(* Logix 5000 project; controller NWGG 1756-L72 rev 35.12; software revision 35.00; part 12 of 19 *)
(* tags used below, declared in another part *)
   _101_FEED_AUGER_PIT_101_HM : HOUR_METER;
   _101M : ALIAS FOR O25[9].3;
   _101Y : ALIAS FOR I25[1].3;
   _102_EXPLORE_TANK_41_RECEIVING_LEG_HM : HOUR_METER;
   _102M : ALIAS FOR O25[8].9;
   _102Y : ALIAS FOR I25[0].9;
   _103_TANK_42_RECEIVING_LEG_HM : HOUR_METER;
   _103_TANK_42_RECEIVING_LEG_RUNNING : BOOL;
   _103M : ALIAS FOR O25[8].12;
   _106_TANK_17_AUGER_HM : HOUR_METER;
   _106_TANK_17_AUGER_RUNNING : BOOL;
   _106M : ALIAS FOR O25[9].5;
   _107_SOUTH_BELT_HM : HOUR_METER;
   _107_TANKS_1THRU7_SOUTH_RUNNING : BOOL;
   _107M : ALIAS FOR O25[9].12;
   _108_CENTER_BELT_HM : HOUR_METER;
   _108_CENTER_BELT_RUNNING : BOOL;
   _109_NORTH_BELT_HM : HOUR_METER;
   _109_RAW_RECEIVING_NORTH_BELT_RUNNING : BOOL;
   _110_TANK_16_AUGER_HM : HOUR_METER;
   _110_TANK_16_AUGER_RUNNING : BOOL;
   _111_TANK_17_AUGER_HM : HOUR_METER;
   _111Y : ALIAS FOR I25[1].0;
   _113_HIGHROLLER_TANKS_11TO15_HM : HOUR_METER;
   _113_HIGHROLLER_TANKS_11TO15_RUNNING : BOOL;
   _113_TO_BC1 : ALIAS FOR O25[11].9;
   _113_TO_BC9 : ALIAS FOR O25[11].8;
   _114_TANKS_1THRU7_NORTH_HM : HOUR_METER;
   _114_TANKS_1THRU7_NORTH_RUNNING : BOOL;
   _116_DRAG_16_HM : HOUR_METER;
   _116Y : ALIAS FOR I25[2].10;
   _117_DRAG_17_HM : HOUR_METER;
   _117Y : ALIAS FOR I25[2].8;
   _11_TANK_41_42_HIGHROLLER_HM : HOUR_METER;
   _11_TANK_41_42_HIGHROLLER_RUNNING : BOOL;
   _11M : ALIAS FOR O25[9].2;
   _122_RECIEVING_LEG_HM : HOUR_METER;
   _122M : ALIAS FOR O25[9].1;
   _122Y : ALIAS FOR I25[1].1;
   _123_CLEAN_LEG_HM : HOUR_METER;
   _123_CLEAN_LEG_RUNNING : BOOL;
   _124M : ALIAS FOR O25[9].13;
   _125_COLOR_SORTER_LEG_HM : HOUR_METER;
   _126_ASPERATOR : HOUR_METER;
   _128_SCREENINGS_DRAG_HM : HOUR_METER;
   _1_CLEAN_SEED_UPPER_BELT_HM : HOUR_METER;
   _1_CLEAN_SEED_UPPER_BELT_RUNNING : BOOL;
   _1M : ALIAS FOR O25[9].8;
   _25_16_0 : ALIAS FOR N200[10];
   _25_16_1 : ALIAS FOR N200[11];
   _25_16_2 : ALIAS FOR N200[12];
   _25_16_3 : ALIAS FOR N200[13];
   _2M : ALIAS FOR O25[9].15;
   _35_JUMP_LEG_HM : HOUR_METER;
   _35_JUMP_LEG_RUNNING : BOOL;
   _36_TANK_41_AUGER_HM : HOUR_METER;
   _36_VFD_TO : ALIAS FOR N180[0];
   _36M : ALIAS FOR O25[8].0;
   _36Y : ALIAS FOR I25[0].0;
   _3_LOWER_TANK_CONVAYOR_24TO26_HM : HOUR_METER;
   _3_LOWER_TANK_CONVAYOR_24TO26_RUNNING : BOOL;
   _3_TO_BC5_S : ALIAS FOR O25[11].12;
   _3_TO_BC6_S : ALIAS FOR O25[11].13;
   _42_LOWER_SCREENINGS_DRAG_HM : HOUR_METER;
   _42M : ALIAS FOR O25[11].1;
   _42Y : ALIAS FOR I25[3].1;
   _43_SCREENINGS_LEG_HM : HOUR_METER;
   _43_SCREENINGS_LEG_RUNNING : BOOL;
   _45M : ALIAS FOR O25[8].7;
   _46M : ALIAS FOR O25[8].8;
   _47M : ALIAS FOR O25[9].10;
   _48_CIMBRIA_HM : HOUR_METER;
   _48_VFD_TO : ALIAS FOR N180[2];
   _48M : ALIAS FOR O25[8].3;
   _48Y : ALIAS FOR I25[0].3;
   _49M : ALIAS FOR O25[9].9;
   _4_LOWER_TANK_CONVAYOR_21TO23_HM : HOUR_METER;
   _4_LOWER_TANK_CONVAYOR_21TO23_RUNNING : BOOL;
   _4_TO_BC5_S : ALIAS FOR O25[11].10;
   _4_TO_BC6_S : ALIAS FOR O25[11].11;
   _50M : ALIAS FOR O25[8].14;
   _51_INDENT_HM : HOUR_METER;
   _51_VFD_TO : ALIAS FOR N180[3];
   _51M : ALIAS FOR O25[8].4;
   _51Y : ALIAS FOR I25[0].4;
   _52M : ALIAS FOR O25[8].6;
   _53_VFD_TO : ALIAS FOR N180[1];
   _53M : ALIAS FOR O25[8].2;
   _54M : ALIAS FOR O25[11].3;
   _55M : ALIAS FOR O25[8].1;
   _56M : ALIAS FOR O25[11].2;
   _57M : ALIAS FOR O25[9].6;
   _5_LOWER_CROSS_BELT_HM : HOUR_METER;
   _5Y : ALIAS FOR I25[2].2;
   _701_TRUCK_REVERSING_BELT_HM : HOUR_METER;
   _701_TRUCK_REVERSING_BELT_RUNNING : BOOL;
   _702_CLEAN_JUMP_BELT_HM : HOUR_METER;
   _702Y : ALIAS FOR I25[1].4;
   _703_TREATER_JUMP_BELT_HM : HOUR_METER;
   _703_TREATER_JUMP_BELT_RUNNING : BOOL;
   _9_TREATER_CONVAYOR_HM : HOUR_METER;
   _9_TREATER_CONVAYOR_RUNNING : BOOL;
   ALARM_HORN : ALIAS FOR O25[11].15;
   ALRM_LIGHT : ALIAS FOR O25[11].14;
   Beta : BOOL;
   CLR_SORT_ASP_DELAY : TIMER;
   CLR_SORT_ASPBLR_DELAY : TIMER;
   CLR_SORT_LEG_DELAY : TIMER;
   CLR_SORT_LEG_SPD10 : ALIAS FOR Local:0:I.Data.3;
   CLR_SORT_LEG_SPD20 : ALIAS FOR Local:0:I.Data.4;
   Consumed : DINT;
   hCLR_SORT_LEG_SPD10 : BOOL;
   hCLR_SORT_LEG_SPD20 : BOOL;
   hCLR_SORT_STB : BOOL;
   hCLR_SORT_STRT : BOOL;
   hN_RECVING_PIT_GATE_CLSPB : BOOL;
   hN_RECVING_PIT_GATE_OPNPB : BOOL;
   hSURGE_BIN_HI : BOOL;
   hSURGE_BIN_LO : BOOL;
   I24 : INT[32];
   I25 : INT[32];
   MTR_125_RUNNING : ALIAS FOR Local:0:I.Data.11;
   MTR_125MB : ALIAS FOR Local:5:O.Data.0;
   MTR_126_RUNNING : ALIAS FOR Local:0:I.Data.6;
   MTR_126M : ALIAS FOR Local:5:O.Data.1;
   MTR_126MB : BOOL;
   MTR_127_RUNNING : ALIAS FOR Local:0:I.Data.7;
   MTR_127M : ALIAS FOR Local:5:O.Data.2;
   MTR_127MB : BOOL;
   MTR_128_RUNNING : ALIAS FOR Local:0:I.Data.5;
   MTR_128M : ALIAS FOR Local:5:O.Data.3;
   MTR_128MB : BOOL;
   N180 : DINT[68];
   N190 : DINT[68];
   N27 : DINT[50];
   N_RECVING_PIT_GATE_AUTO : ALIAS FOR Local:0:I.Data.2;
   N_RECVING_PIT_GATE_CLOSE : ALIAS FOR Local:5:O.Data.5;
   N_RECVING_PIT_GATE_OPEN : ALIAS FOR Local:5:O.Data.4;
   O24 : INT[32];
   O25 : INT[32];
   O25_012_Bit00 : ALIAS FOR O25[12].0;
   O25_012_Bit01 : ALIAS FOR O25[12].1;
   O25_012_Bit02 : ALIAS FOR O25[12].2;
   O25_012_Bit03 : ALIAS FOR O25[12].3;
   O25_012_Bit04 : ALIAS FOR O25[12].4;
   O25_012_Bit05 : ALIAS FOR O25[12].5;
   O25_012_Bit06 : ALIAS FOR O25[12].6;
   O25_012_Bit07 : ALIAS FOR O25[12].7;
   O25_012_Bit08 : ALIAS FOR O25[12].8;
   O25_012_Bit09 : ALIAS FOR O25[12].9;
   O25_012_Bit10 : ALIAS FOR O25[12].10;
   O25_012_Bit11 : ALIAS FOR O25[12].11;
   O25_012_Bit12 : ALIAS FOR O25[12].12;
   O25_012_Bit13 : ALIAS FOR O25[12].13;
   O25_012_Bit14 : ALIAS FOR O25[12].14;
   output_Bit : BOOL;
   Output_Bit_2 : BOOL;
   Rack24_1_Mode : BOOL;
   SURGE_BIN_HI : ALIAS FOR Local:0:I.Data.0;
   SURGE_BIN_LO : ALIAS FOR Local:0:I.Data.1;
(* MainProgram, continued *)

ROUTINE Dev_O25_11   (* ladder *)
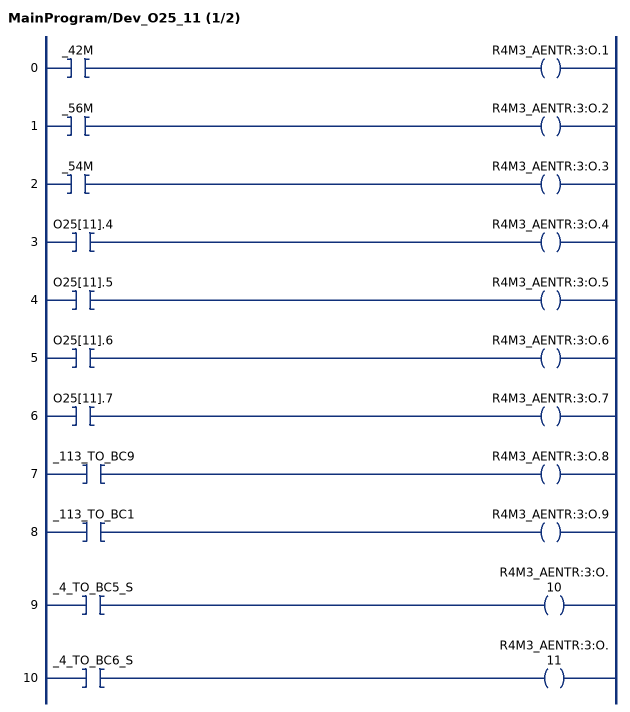
   0: XIC(_42M)OTE(R4M3_AENTR:3:O.1);
   1: XIC(_56M)OTE(R4M3_AENTR:3:O.2);
   2: XIC(_54M)OTE(R4M3_AENTR:3:O.3);
   3: XIC(O25[11].4)OTE(R4M3_AENTR:3:O.4);
   4: XIC(O25[11].5)OTE(R4M3_AENTR:3:O.5);
   5: XIC(O25[11].6)OTE(R4M3_AENTR:3:O.6);
   6: XIC(O25[11].7)OTE(R4M3_AENTR:3:O.7);
   7: XIC(_113_TO_BC9)OTE(R4M3_AENTR:3:O.8);
   8: XIC(_113_TO_BC1)OTE(R4M3_AENTR:3:O.9);
   9: XIC(_4_TO_BC5_S)OTE(R4M3_AENTR:3:O.10);
   10: XIC(_4_TO_BC6_S)OTE(R4M3_AENTR:3:O.11);
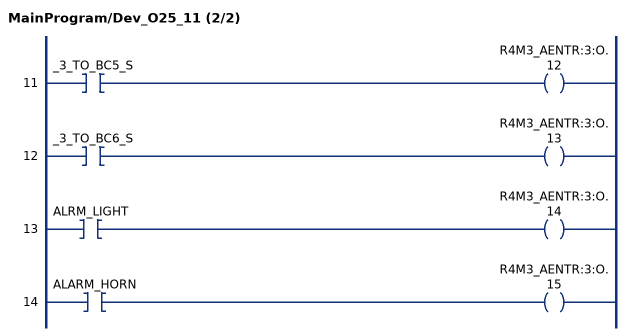
   11: XIC(_3_TO_BC5_S)OTE(R4M3_AENTR:3:O.12);
   12: XIC(_3_TO_BC6_S)OTE(R4M3_AENTR:3:O.13);
   13: XIC(ALRM_LIGHT)OTE(R4M3_AENTR:3:O.14);
   14: XIC(ALARM_HORN)OTE(R4M3_AENTR:3:O.15);
END_ROUTINE

ROUTINE Dev_O25_12   (* ladder *)
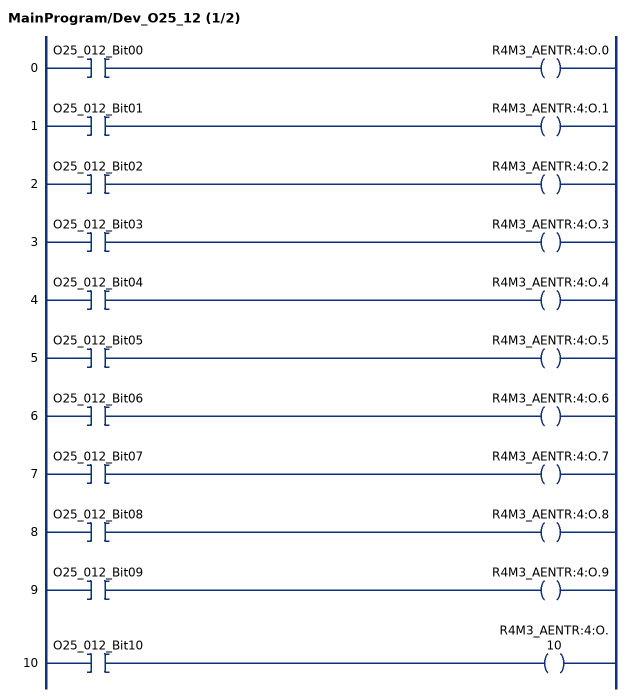
   0: XIC(O25_012_Bit00)OTE(R4M3_AENTR:4:O.0);
   1: XIC(O25_012_Bit01)OTE(R4M3_AENTR:4:O.1);
   2: XIC(O25_012_Bit02)OTE(R4M3_AENTR:4:O.2);
   3: XIC(O25_012_Bit03)OTE(R4M3_AENTR:4:O.3);
   4: XIC(O25_012_Bit04)OTE(R4M3_AENTR:4:O.4);
   5: XIC(O25_012_Bit05)OTE(R4M3_AENTR:4:O.5);
   6: XIC(O25_012_Bit06)OTE(R4M3_AENTR:4:O.6);
   7: XIC(O25_012_Bit07)OTE(R4M3_AENTR:4:O.7);
   8: XIC(O25_012_Bit08)OTE(R4M3_AENTR:4:O.8);
   9: XIC(O25_012_Bit09)OTE(R4M3_AENTR:4:O.9);
   10: XIC(O25_012_Bit10)OTE(R4M3_AENTR:4:O.10);
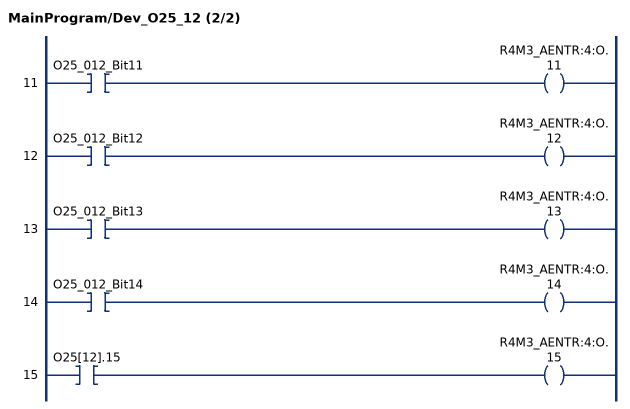
   11: XIC(O25_012_Bit11)OTE(R4M3_AENTR:4:O.11);
   12: XIC(O25_012_Bit12)OTE(R4M3_AENTR:4:O.12);
   13: XIC(O25_012_Bit13)OTE(R4M3_AENTR:4:O.13);
   14: XIC(O25_012_Bit14)OTE(R4M3_AENTR:4:O.14);
   15: XIC(O25[12].15)OTE(R4M3_AENTR:4:O.15);
END_ROUTINE

ROUTINE Dev_O25_8   (* ladder *)
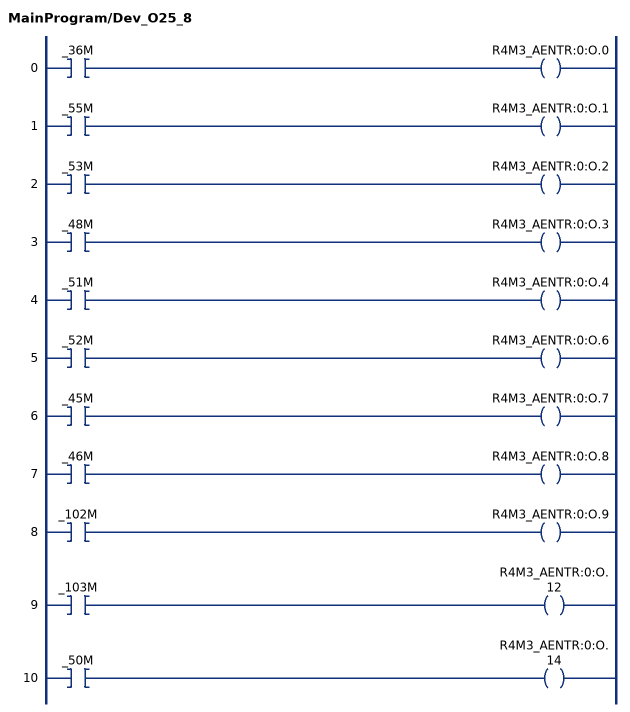
   0: XIC(_36M)OTE(R4M3_AENTR:0:O.0);
   1: XIC(_55M)OTE(R4M3_AENTR:0:O.1);
   2: XIC(_53M)OTE(R4M3_AENTR:0:O.2);
   3: XIC(_48M)OTE(R4M3_AENTR:0:O.3);
   4: XIC(_51M)OTE(R4M3_AENTR:0:O.4);
   5: XIC(_52M)OTE(R4M3_AENTR:0:O.6);
   6: XIC(_45M)OTE(R4M3_AENTR:0:O.7);
   7: XIC(_46M)OTE(R4M3_AENTR:0:O.8);
   8: XIC(_102M)OTE(R4M3_AENTR:0:O.9);
   9: XIC(_103M)OTE(R4M3_AENTR:0:O.12);
   10: XIC(_50M)OTE(R4M3_AENTR:0:O.14);
END_ROUTINE

ROUTINE Dev_O25_9   (* ladder *)
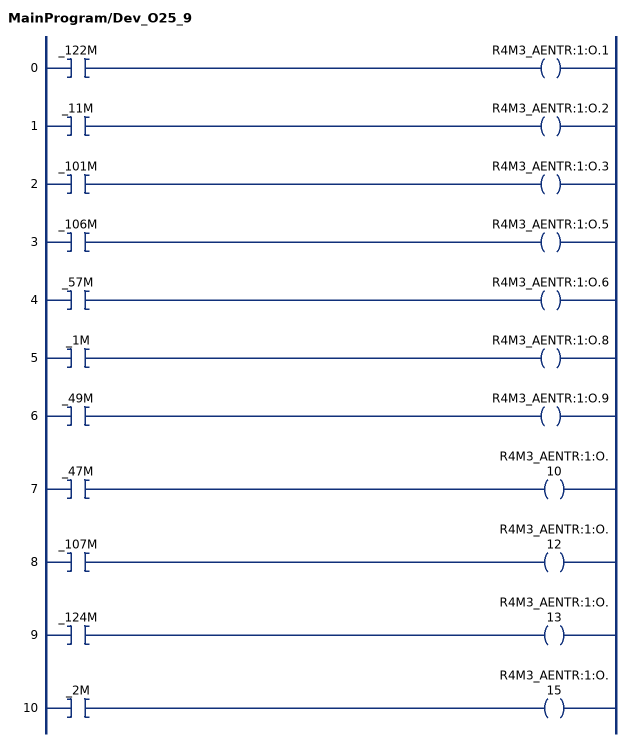
   0: XIC(_122M)OTE(R4M3_AENTR:1:O.1);
   1: XIC(_11M)OTE(R4M3_AENTR:1:O.2);
   2: XIC(_101M)OTE(R4M3_AENTR:1:O.3);
   3: XIC(_106M)OTE(R4M3_AENTR:1:O.5);
   4: XIC(_57M)OTE(R4M3_AENTR:1:O.6);
   5: XIC(_1M)OTE(R4M3_AENTR:1:O.8);
   6: XIC(_49M)OTE(R4M3_AENTR:1:O.9);
   7: XIC(_47M)OTE(R4M3_AENTR:1:O.10);
   8: XIC(_107M)OTE(R4M3_AENTR:1:O.12);
   9: XIC(_124M)OTE(R4M3_AENTR:1:O.13);
   10: XIC(_2M)OTE(R4M3_AENTR:1:O.15);
END_ROUTINE

ROUTINE Disp   (* ladder *)
END_ROUTINE

ROUTINE HOUR_METERS   (* ladder *)
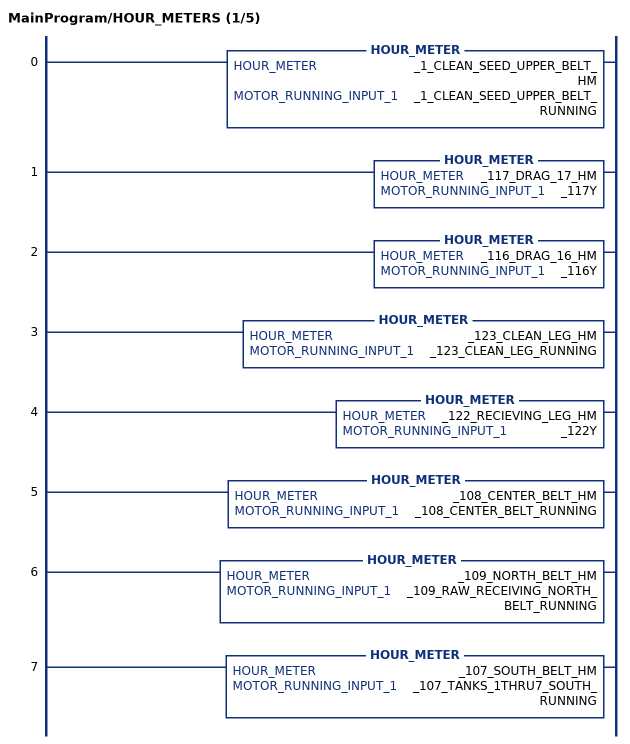
   0: HOUR_METER(_1_CLEAN_SEED_UPPER_BELT_HM,_1_CLEAN_SEED_UPPER_BELT_RUNNING);
   1: HOUR_METER(_117_DRAG_17_HM,_117Y);
   2: HOUR_METER(_116_DRAG_16_HM,_116Y);
   3: HOUR_METER(_123_CLEAN_LEG_HM,_123_CLEAN_LEG_RUNNING);
   4: HOUR_METER(_122_RECIEVING_LEG_HM,_122Y);
   5: HOUR_METER(_108_CENTER_BELT_HM,_108_CENTER_BELT_RUNNING);
   6: HOUR_METER(_109_NORTH_BELT_HM,_109_RAW_RECEIVING_NORTH_BELT_RUNNING);
   7: HOUR_METER(_107_SOUTH_BELT_HM,_107_TANKS_1THRU7_SOUTH_RUNNING);
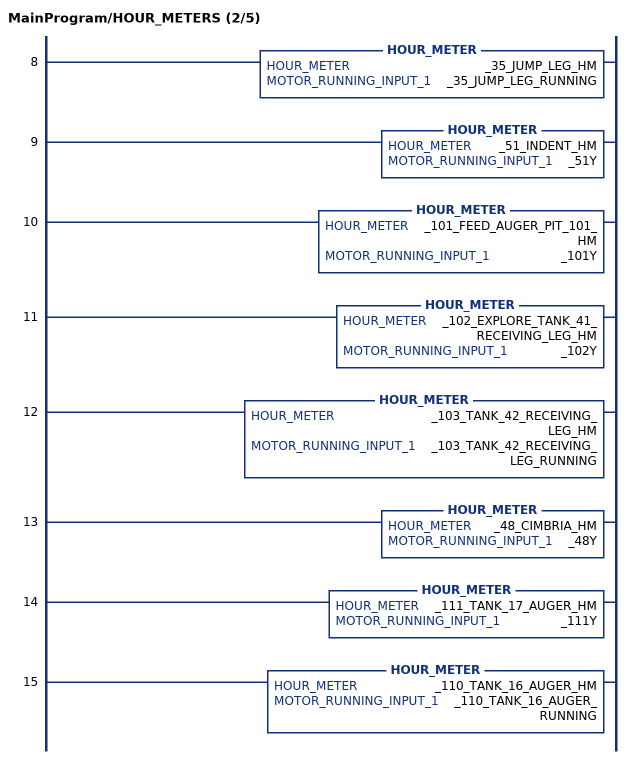
   8: HOUR_METER(_35_JUMP_LEG_HM,_35_JUMP_LEG_RUNNING);
   9: HOUR_METER(_51_INDENT_HM,_51Y);
   10: HOUR_METER(_101_FEED_AUGER_PIT_101_HM,_101Y);
   11: HOUR_METER(_102_EXPLORE_TANK_41_RECEIVING_LEG_HM,_102Y);
   12: HOUR_METER(_103_TANK_42_RECEIVING_LEG_HM,_103_TANK_42_RECEIVING_LEG_RUNNING);
   13: HOUR_METER(_48_CIMBRIA_HM,_48Y);
   14: HOUR_METER(_111_TANK_17_AUGER_HM,_111Y);
   15: HOUR_METER(_110_TANK_16_AUGER_HM,_110_TANK_16_AUGER_RUNNING);
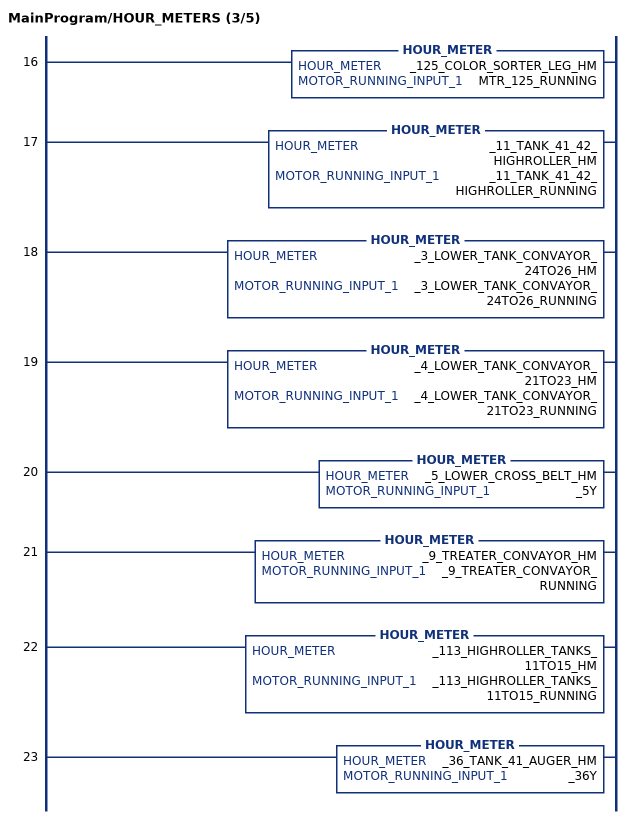
   16: HOUR_METER(_125_COLOR_SORTER_LEG_HM,MTR_125_RUNNING);
   17: HOUR_METER(_11_TANK_41_42_HIGHROLLER_HM,_11_TANK_41_42_HIGHROLLER_RUNNING);
   18: HOUR_METER(_3_LOWER_TANK_CONVAYOR_24TO26_HM,_3_LOWER_TANK_CONVAYOR_24TO26_RUNNING);
   19: HOUR_METER(_4_LOWER_TANK_CONVAYOR_21TO23_HM,_4_LOWER_TANK_CONVAYOR_21TO23_RUNNING);
   20: HOUR_METER(_5_LOWER_CROSS_BELT_HM,_5Y);
   21: HOUR_METER(_9_TREATER_CONVAYOR_HM,_9_TREATER_CONVAYOR_RUNNING);
   22: HOUR_METER(_113_HIGHROLLER_TANKS_11TO15_HM,_113_HIGHROLLER_TANKS_11TO15_RUNNING);
   23: HOUR_METER(_36_TANK_41_AUGER_HM,_36Y);
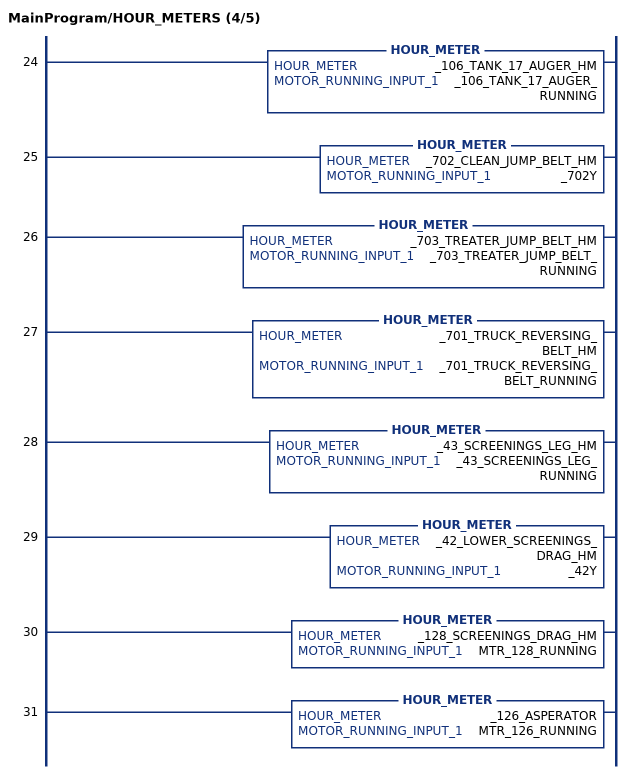
   24: HOUR_METER(_106_TANK_17_AUGER_HM,_106_TANK_17_AUGER_RUNNING);
   25: HOUR_METER(_702_CLEAN_JUMP_BELT_HM,_702Y);
   26: HOUR_METER(_703_TREATER_JUMP_BELT_HM,_703_TREATER_JUMP_BELT_RUNNING);
   27: HOUR_METER(_701_TRUCK_REVERSING_BELT_HM,_701_TRUCK_REVERSING_BELT_RUNNING);
   28: HOUR_METER(_43_SCREENINGS_LEG_HM,_43_SCREENINGS_LEG_RUNNING);
   29: HOUR_METER(_42_LOWER_SCREENINGS_DRAG_HM,_42Y);
   30: HOUR_METER(_128_SCREENINGS_DRAG_HM,MTR_128_RUNNING);
   31: HOUR_METER(_126_ASPERATOR,MTR_126_RUNNING);
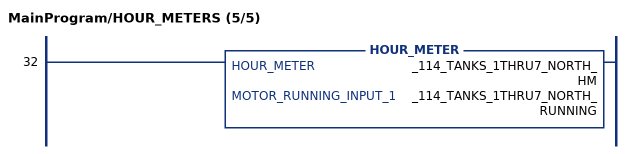
   32: HOUR_METER(_114_TANKS_1THRU7_NORTH_HM,_114_TANKS_1THRU7_NORTH_RUNNING);
END_ROUTINE

ROUTINE MainRoutine   (* ladder *)
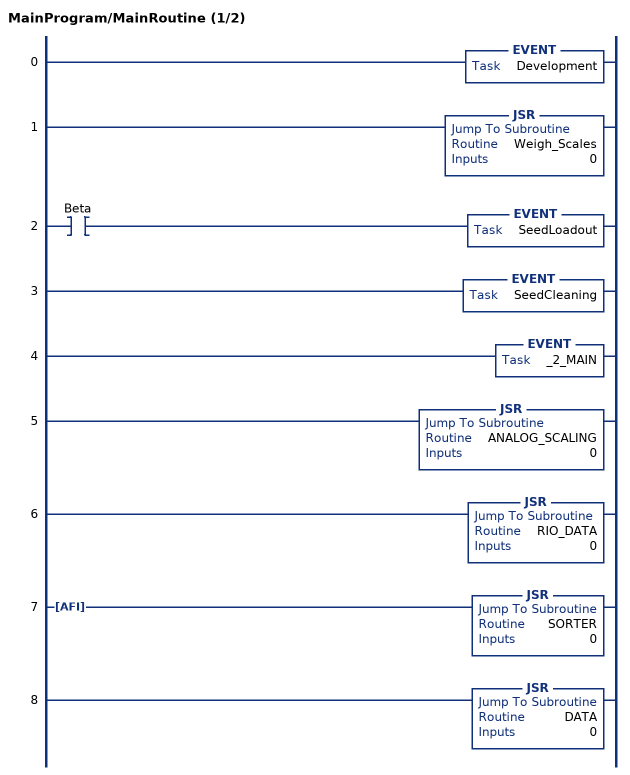
   0: EVENT(Development);
   1: JSR(Weigh_Scales,0);
   2: XIC(Beta)EVENT(SeedLoadout);
   3: EVENT(SeedCleaning);
   4: EVENT(_2_MAIN);
   5: JSR(ANALOG_SCALING,0);
   6: JSR(RIO_DATA,0);
   7: AFI()JSR(SORTER,0);
   8: JSR(DATA,0);
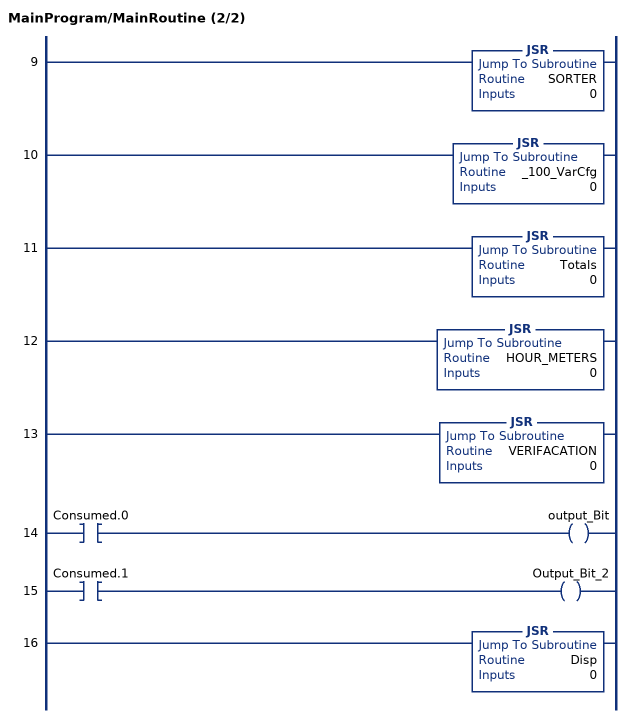
   9: JSR(SORTER,0);
   10: JSR(_100_VarCfg,0);
   11: JSR(Totals,0);
   12: JSR(HOUR_METERS,0);
   13: JSR(VERIFACATION,0);
   14: XIC(Consumed.0)OTE(output_Bit);
   15: XIC(Consumed.1)OTE(Output_Bit_2);
   16: JSR(Disp,0);
END_ROUTINE

ROUTINE RIO_DATA   (* ladder *)
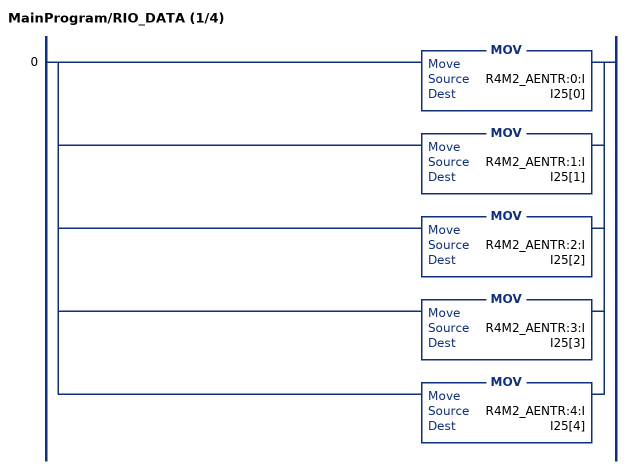
   0: [MOV(R4M2_AENTR:0:I,I25[0]) ,MOV(R4M2_AENTR:1:I,I25[1]) ,MOV(R4M2_AENTR:2:I,I25[2]) ,MOV(R4M2_AENTR:3:I,I25[3]) ,MOV(R4M2_AENTR:4:I,I25[4]) ];
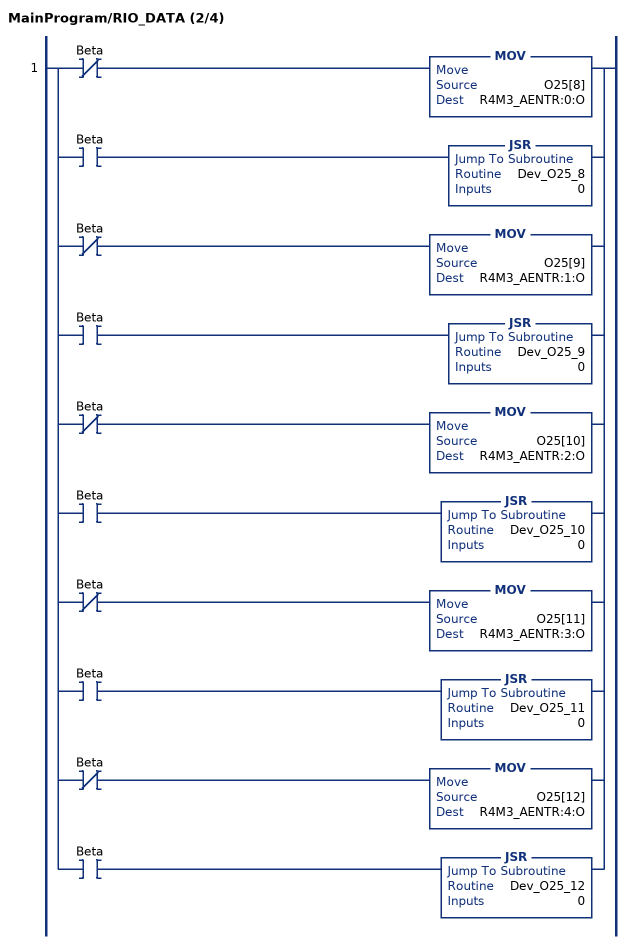
   1: [XIO(Beta) MOV(O25[8],R4M3_AENTR:0:O) ,XIC(Beta) JSR(Dev_O25_8,0) ,XIO(Beta) MOV(O25[9],R4M3_AENTR:1:O) ,XIC(Beta) JSR(Dev_O25_9,0) ,XIO(Beta) MOV(O25[10],R4M3_AENTR:2:O) ,XIC(Beta) JSR(Dev_O25_10,0) ,XIO(Beta) MOV(O25[11],R4M3_AENTR:3:O) ,XIC(Beta) JSR(Dev_O25_11,0) ,XIO(Beta) MOV(O25[12],R4M3_AENTR:4:O) ,XIC(Beta) JSR(Dev_O25_12,0) ];
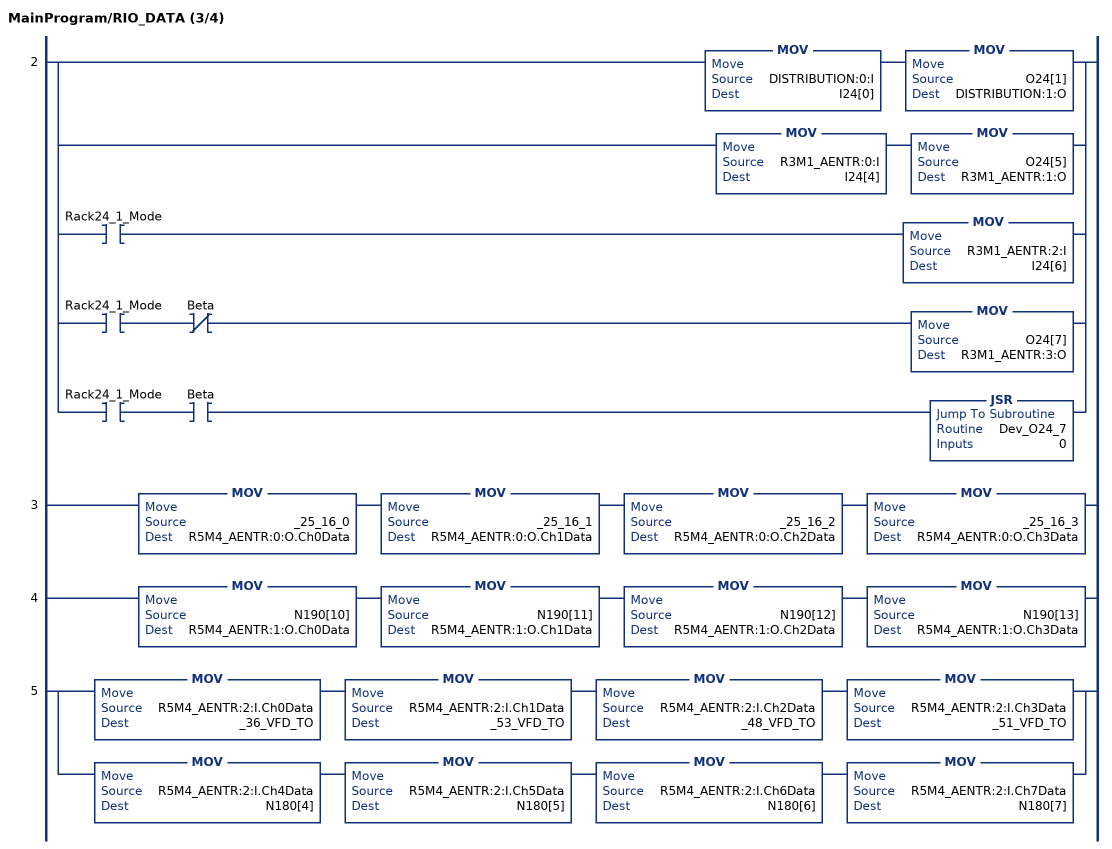
   2: [MOV(DISTRIBUTION:0:I,I24[0]) MOV(O24[1],DISTRIBUTION:1:O) ,MOV(R3M1_AENTR:0:I,I24[4]) MOV(O24[5],R3M1_AENTR:1:O) ,XIC(Rack24_1_Mode) MOV(R3M1_AENTR:2:I,I24[6]) ,XIC(Rack24_1_Mode) XIO(Beta) MOV(O24[7],R3M1_AENTR:3:O) ,XIC(Rack24_1_Mode) XIC(Beta) JSR(Dev_O24_7,0) ];
   3: MOV(_25_16_0,R5M4_AENTR:0:O.Ch0Data)MOV(_25_16_1,R5M4_AENTR:0:O.Ch1Data)MOV(_25_16_2,R5M4_AENTR:0:O.Ch2Data)MOV(_25_16_3,R5M4_AENTR:0:O.Ch3Data);
   4: MOV(N190[10],R5M4_AENTR:1:O.Ch0Data)MOV(N190[11],R5M4_AENTR:1:O.Ch1Data)MOV(N190[12],R5M4_AENTR:1:O.Ch2Data)MOV(N190[13],R5M4_AENTR:1:O.Ch3Data);
   5: [MOV(R5M4_AENTR:2:I.Ch0Data,_36_VFD_TO) MOV(R5M4_AENTR:2:I.Ch1Data,_53_VFD_TO) MOV(R5M4_AENTR:2:I.Ch2Data,_48_VFD_TO) MOV(R5M4_AENTR:2:I.Ch3Data,_51_VFD_TO) ,MOV(R5M4_AENTR:2:I.Ch4Data,N180[4]) MOV(R5M4_AENTR:2:I.Ch5Data,N180[5]) MOV(R5M4_AENTR:2:I.Ch6Data,N180[6]) MOV(R5M4_AENTR:2:I.Ch7Data,N180[7]) ];
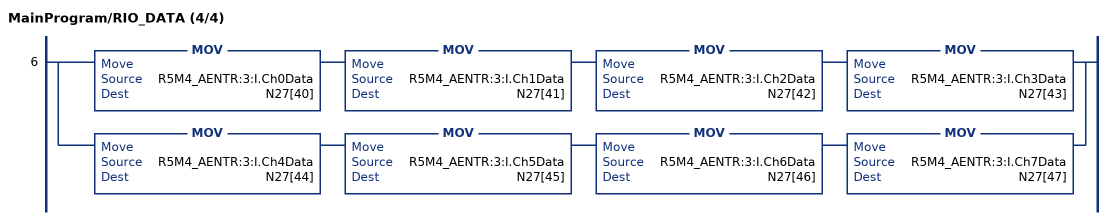
   6: [MOV(R5M4_AENTR:3:I.Ch0Data,N27[40]) MOV(R5M4_AENTR:3:I.Ch1Data,N27[41]) MOV(R5M4_AENTR:3:I.Ch2Data,N27[42]) MOV(R5M4_AENTR:3:I.Ch3Data,N27[43]) ,MOV(R5M4_AENTR:3:I.Ch4Data,N27[44]) MOV(R5M4_AENTR:3:I.Ch5Data,N27[45]) MOV(R5M4_AENTR:3:I.Ch6Data,N27[46]) MOV(R5M4_AENTR:3:I.Ch7Data,N27[47]) ];
END_ROUTINE

ROUTINE SORTER   (* ladder *)
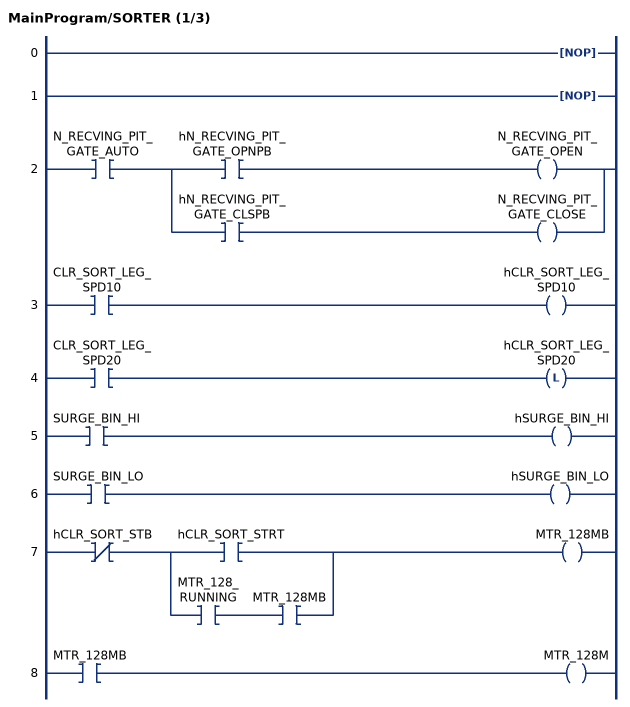
   0: NOP();
   1: NOP();
   2: XIC(N_RECVING_PIT_GATE_AUTO)[XIC(hN_RECVING_PIT_GATE_OPNPB) OTE(N_RECVING_PIT_GATE_OPEN) ,XIC(hN_RECVING_PIT_GATE_CLSPB) OTE(N_RECVING_PIT_GATE_CLOSE) ];
   3: XIC(CLR_SORT_LEG_SPD10)OTE(hCLR_SORT_LEG_SPD10);
   4: XIC(CLR_SORT_LEG_SPD20)OTL(hCLR_SORT_LEG_SPD20);
   5: XIC(SURGE_BIN_HI)OTE(hSURGE_BIN_HI);
   6: XIC(SURGE_BIN_LO)OTE(hSURGE_BIN_LO);
   7: XIO(hCLR_SORT_STB)[XIC(hCLR_SORT_STRT) ,XIC(MTR_128_RUNNING) XIC(MTR_128MB) ]OTE(MTR_128MB);
   8: XIC(MTR_128MB)OTE(MTR_128M);
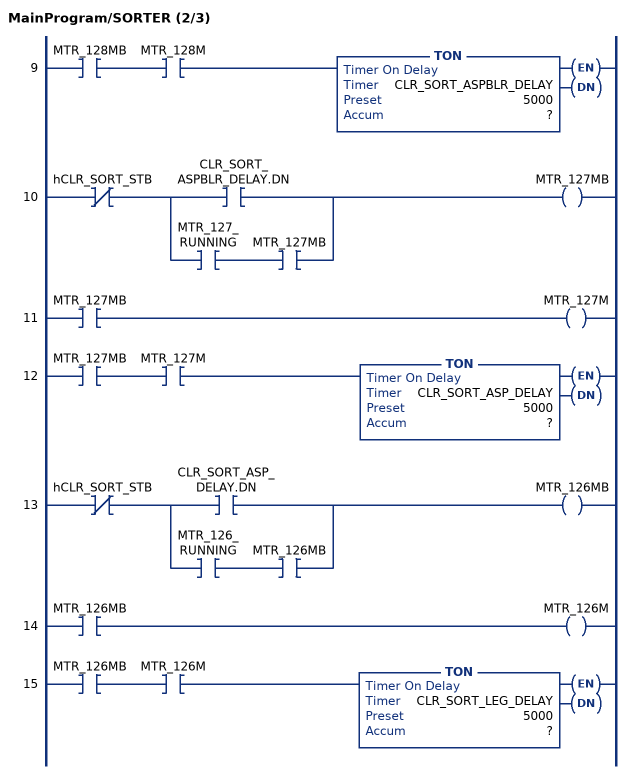
   9: XIC(MTR_128MB)XIC(MTR_128M)TON(CLR_SORT_ASPBLR_DELAY,?,?);
   10: XIO(hCLR_SORT_STB)[XIC(CLR_SORT_ASPBLR_DELAY.DN) ,XIC(MTR_127_RUNNING) XIC(MTR_127MB) ]OTE(MTR_127MB);
   11: XIC(MTR_127MB)OTE(MTR_127M);
   12: XIC(MTR_127MB)XIC(MTR_127M)TON(CLR_SORT_ASP_DELAY,?,?);
   13: XIO(hCLR_SORT_STB)[XIC(CLR_SORT_ASP_DELAY.DN) ,XIC(MTR_126_RUNNING) XIC(MTR_126MB) ]OTE(MTR_126MB);
   14: XIC(MTR_126MB)OTE(MTR_126M);
   15: XIC(MTR_126MB)XIC(MTR_126M)TON(CLR_SORT_LEG_DELAY,?,?);
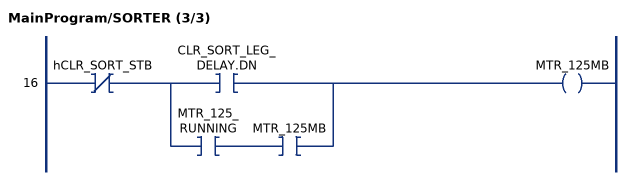
   16: XIO(hCLR_SORT_STB)[XIC(CLR_SORT_LEG_DELAY.DN) ,XIC(MTR_125_RUNNING) XIC(MTR_125MB) ]OTE(MTR_125MB);
END_ROUTINE
